screen "RIO 02 Digital Inputs" 1280x800, template "Template"
   on GenerateScreen: "TitleUpdater"()
   TextField "Text field_37" at 16,52 size 476x26; Text 'RIO #2 (Remote Inputs & Outputs Panel No. 2)'
   TextField "Text field_38" at 16,122 size 55x22; Text 'I15.0'
   TextField "Text field_39" at 16,157 size 55x22; Text 'I15.1'
   TextField "Text field_40" at 16,193 size 55x22; Text 'I15.2'
   TextField "Text field_41" at 16,229 size 55x22; Text 'I15.3'
   TextField "Text field_42" at 16,265 size 55x22; Text 'I15.4'
   TextField "Text field_43" at 16,301 size 55x22; Text 'I15.5'
   TextField "Text field_44" at 16,337 size 55x22; Text 'I15.6'
   TextField "Text field_45" at 16,373 size 55x22; Text 'I15.7'
   Circle "Circle_33" at 76,123 size 20x20
      Appearance <- "Tank 2P GTT Isolation Valve Feedback - Opened"
   Circle "Circle_34" at 76,158 size 20x20
      Appearance <- "Tank 2P GTT Isolation Valve Feedback - Closed"
   Circle "Circle_35" at 76,194 size 20x20
      Appearance <- "Tank 2P Tank Vent Valve 1 Feedback - Opened"
   Circle "Circle_36" at 76,230 size 20x20
      Appearance <- "Tank 2P Tank Vent Valve 1 Feedback - Closed"
   Circle "Circle_37" at 76,265 size 20x20
      Appearance <- "Tank 2P Tank Vent Valve 2 Feedback - Opened"
   Circle "Circle_38" at 76,301 size 20x20
      Appearance <- "Tank 2P Tank Vent Valve 2 Feedback - Closed"
   Circle "Circle_39" at 76,337 size 20x20
      Appearance <- "RIO2_SPR_DI_15_6"
   Circle "Circle_40" at 76,373 size 20x20
      Appearance <- "RIO2_SPR_DI_15_7"
   TextField "Text field_46" at 33,90 size 49x26; Text 'I0'
   TextField "Text field_47" at 16,441 size 55x22; Text 'I18.0'
   TextField "Text field_48" at 16,476 size 55x22; Text 'I18.1'
   TextField "Text field_49" at 16,512 size 55x22; Text 'I18.2'
   TextField "Text field_50" at 16,548 size 55x22; Text 'I18.3'
   TextField "Text field_51" at 16,584 size 55x22; Text 'I18.4'
   TextField "Text field_52" at 16,620 size 55x22; Text 'I18.5'
   TextField "Text field_53" at 16,656 size 55x22; Text 'I18.6'
   TextField "Text field_54" at 16,692 size 55x22; Text 'I18.7'
   Circle "Circle_41" at 76,442 size 20x20
      Appearance <- "Tank 2S GTT Isolation Valve Feedback - Opened"
   Circle "Circle_42" at 76,477 size 20x20
      Appearance <- "Tank 2S GTT Isolation Valve Feedback - Closed"
   Circle "Circle_43" at 76,513 size 20x20
      Appearance <- "Tank 2S Tank Vent Valve 1 Feedback - Opened"
   Circle "Circle_44" at 76,549 size 20x20
      Appearance <- "Tank 2S Tank Vent Valve 1 Feedback - Closed"
   Circle "Circle_45" at 76,585 size 20x20
      Appearance <- "Tank 2S Tank Vent Valve 2 Feedback - Opened"
   Circle "Circle_46" at 76,621 size 20x20
      Appearance <- "Tank 2S Tank Vent Valve 2 Feedback - Closed"
   Circle "Circle_47" at 76,657 size 20x20
      Appearance <- "RIO2_SPR_DI_18_6"
   Circle "Circle_48" at 76,693 size 20x20
      Appearance <- "RIO2_SPR_DI_18_7"
   TextField "Text field_55" at 33,409 size 49x26; Text 'I1'
   TextField "Text field_56" at 548,122 size 55x22; Text 'I21.0'
   TextField "Text field_57" at 548,157 size 55x22; Text 'I21.1'
   TextField "Text field_58" at 548,193 size 55x22; Text 'I21.2'
   TextField "Text field_59" at 548,229 size 55x22; Text 'I21.3'
   TextField "Text field_60" at 548,265 size 55x22; Text 'I21.4'
   TextField "Text field_61" at 548,301 size 55x22; Text 'I21.5'
   TextField "Text field_62" at 548,337 size 55x22; Text 'I21.6'
   TextField "Text field_63" at 548,373 size 55x22; Text 'I21.7'
   Circle "Circle_49" at 608,122 size 20x20
      Appearance <- "Tank 2P BWT Level High High Switch"
   Circle "Circle_50" at 608,157 size 20x20
      Appearance <- "RIO2 Tanks Pressure Switch Hi Hi"
   Circle "Circle_51" at 608,193 size 20x20
      Appearance <- "Tank 2S BWT Level High High Switch"
   Circle "Circle_52" at 608,229 size 20x20
      Appearance <- "RIO2_SPR_DI_21_3"
   Circle "Circle_53" at 608,265 size 20x20
      Appearance <- "RIO2_SPR_DI_21_4"
   Circle "Circle_54" at 608,301 size 20x20
      Appearance <- "RIO2_SPR_DI_21_5"
   Circle "Circle_55" at 608,337 size 20x20
      Appearance <- "RIO2_SPR_DI_21_6"
   Circle "Circle_56" at 608,373 size 20x20
      Appearance <- "RIO2_SPR_DI_21_7"
   TextField "Text field_64" at 570,90 size 49x26; Text 'I2'
   Button "HmiScreenItemData_1" at 1,1 size 150x43; TextOn 'Back'; TextOff 'Commissioning'
      on Release: ActivateScreen("Commissioning Main Page", 0)
   TextField "Text field_107" at 105,114 size 382x38; Text 'Tank 2P GTT Isolation Valve Feedback - Opened CV422'
   TextField "Text field_108" at 105,149 size 374x38; Text 'Tank 2P GTT Isolation Valve Feedback - Closed CV422'
   TextField "Text field_109" at 105,184 size 371x38; Text 'Tank 2P Tank Vent Valve 1 Feedback - Opened CV441-2P1'
   TextField "Text field_110" at 105,220 size 363x38; Text 'Tank 2P Tank Vent Valve 1 Feedback - Closed CV441-2P1'
   TextField "Text field_111" at 105,255 size 371x38; Text 'Tank 2P Tank Vent Valve 2 Feedback - Opened CV441-2P2'
   TextField "Text field_112" at 105,291 size 363x38; Text 'Tank 2P Tank Vent Valve 2 Feedback - Closed CV441-2P2'
   TextField "Text field_113" at 104,328 size 100x21; Text 'Spare Input'
   TextField "Text field_114" at 104,365 size 100x21; Text 'Spare Input'
   TextField "Text field_116" at 102,429 size 382x38; Text 'Tank 2S GTT Isolation Valve Feedback - Opened CV421-2S'
   TextField "Text field_117" at 102,465 size 374x38; Text 'Tank 2S GTT Isolation Valve Feedback - Closed CV421-2S'
   TextField "Text field_118" at 102,501 size 371x38; Text 'Tank 2S Tank Vent Valve 1 Feedback - Opened CV440-2SA'
   TextField "Text field_119" at 102,537 size 363x38; Text 'Tank 2S Tank Vent Valve 1 Feedback - Closed CV440-2SA'
   TextField "Text field_120" at 102,573 size 371x38; Text 'Tank 2S Tank Vent Valve 2 Feedback - Opened CV440-2SB'
   TextField "Text field_121" at 102,609 size 363x38; Text 'Tank 2S Tank Vent Valve 2 Feedback - Closed CV440-2SB'
   TextField "Text field_122" at 102,690 size 100x21; Text 'Spare Input'
   TextField "Text field_123" at 636,113 size 294x38; Text 'Tank 2P BWT Level High High Switch LS425-2P'
   TextField "Text field_124" at 636,148 size 270x38; Text 'RIO2 Tanks Pressure Switch Hi Hi PS436-2P/2S'
   TextField "Text field_125" at 636,184 size 294x38; Text 'Tank 2S BWT Level High High Switch LS422-2S'
   TextField "Text field_126" at 636,219 size 100x21; Text 'Spare Input'
   TextField "Text field_127" at 636,255 size 100x21; Text 'Spare Input'
   TextField "Text field_128" at 636,291 size 100x21; Text 'Spare Input'
   TextField "Text field_129" at 636,328 size 100x21; Text 'Spare Input'
   TextField "Text field_130" at 636,366 size 100x21; Text 'Spare Input'
   TextField "Text field_115" at 102,654 size 100x21; Text 'Spare Input'
   AlarmView "Alarm view_1" at 0,777 size 1280x23
   Group "Group" at 455,41 size 373x50
   Button "HmiScreenItemData_8" at 469,45 size 355x40; TextOn 'Back'; TextOff 'Text'
      on Click: "TitleUpdater"()
   TextField "Screen title" at 455,41 size 373x50; Text 'Screen title'

screen "RIO 03 Digital Inputs" 1280x800, template "Template"
   on GenerateScreen: "TitleUpdater"()
   TextField "Text field_37" at 16,52 size 476x26; Text 'RIO #3 (Remote Inputs & Outputs Panel No. 3)'
   TextField "Text field_38" at 16,122 size 55x22; Text 'I27.0'
   TextField "Text field_39" at 16,157 size 55x22; Text 'I27.1'
   TextField "Text field_40" at 16,193 size 55x22; Text 'I27.2'
   TextField "Text field_41" at 16,229 size 55x22; Text 'I27.3'
   TextField "Text field_42" at 16,265 size 55x22; Text 'I27.4'
   TextField "Text field_43" at 16,301 size 55x22; Text 'I27.5'
   TextField "Text field_44" at 16,337 size 55x22; Text 'I27.6'
   TextField "Text field_45" at 16,373 size 55x22; Text 'I27.7'
   Circle "Circle_33" at 76,123 size 20x20
      Appearance <- "Tank 3P GTT Isolation Valve Feedback - Opened"
   Circle "Circle_34" at 76,158 size 20x20
      Appearance <- "Tank 3P GTT Isolation Valve Feedback - Closed"
   Circle "Circle_35" at 76,194 size 20x20
      Appearance <- "Tank 3P Tank Vent Valve 1 Feedback - Opened"
   Circle "Circle_36" at 76,230 size 20x20
      Appearance <- "Tank 3P Tank Vent Valve 1 Feedback - Closed"
   Circle "Circle_37" at 76,265 size 20x20
      Appearance <- "Tank 3P Tank Vent Valve 2 Feedback - Opened"
   Circle "Circle_38" at 76,301 size 20x20
      Appearance <- "Tank 3P Tank Vent Valve 2 Feedback - Closed"
   Circle "Circle_39" at 76,337 size 20x20
      Appearance <- "RIO3_SPR_DI_27_6"
   Circle "Circle_40" at 76,373 size 20x20
      Appearance <- "RIO3_SPR_DI_27_7"
   TextField "Text field_46" at 33,90 size 49x26; Text 'I0'
   TextField "Text field_47" at 16,441 size 55x22; Text 'I30.0'
   TextField "Text field_48" at 16,476 size 55x22; Text 'I30.1'
   TextField "Text field_49" at 16,512 size 55x22; Text 'I30.2'
   TextField "Text field_50" at 16,548 size 55x22; Text 'I30.3'
   TextField "Text field_51" at 16,584 size 55x22; Text 'I30.4'
   TextField "Text field_52" at 16,620 size 55x22; Text 'I30.5'
   TextField "Text field_53" at 16,656 size 55x22; Text 'I30.6'
   TextField "Text field_54" at 16,692 size 55x22; Text 'I30.7'
   Circle "Circle_41" at 76,442 size 20x20
      Appearance <- "Tank 3S GTT Isolation Valve Feedback - Opened"
   Circle "Circle_42" at 76,477 size 20x20
      Appearance <- "Tank 3S GTT Isolation Valve Feedback - Closed"
   Circle "Circle_43" at 76,513 size 20x20
      Appearance <- "Tank 3S Tank Vent Valve 1 Feedback - Opened"
   Circle "Circle_44" at 76,549 size 20x20
      Appearance <- "Tank 3S Tank Vent Valve 1 Feedback - Closed"
   Circle "Circle_45" at 76,585 size 20x20
      Appearance <- "Tank 3S Tank Vent Valve 2 Feedback - Opened"
   Circle "Circle_46" at 76,621 size 20x20
      Appearance <- "Tank 3S Tank Vent Valve 2 Feedback - Closed"
   Circle "Circle_47" at 76,657 size 20x20
      Appearance <- "RIO3_SPR_DI_30_6"
   Circle "Circle_48" at 76,693 size 20x20
      Appearance <- "RIO3_SPR_DI_30_7"
   TextField "Text field_55" at 33,409 size 49x26; Text 'I1'
   TextField "Text field_56" at 548,122 size 55x22; Text 'I33.0'
   TextField "Text field_57" at 548,157 size 55x22; Text 'I33.1'
   TextField "Text field_58" at 548,193 size 55x22; Text 'I33.2'
   TextField "Text field_59" at 548,229 size 55x22; Text 'I33.3'
   TextField "Text field_60" at 548,265 size 55x22; Text 'I33.4'
   TextField "Text field_61" at 548,301 size 55x22; Text 'I33.5'
   TextField "Text field_62" at 548,337 size 55x22; Text 'I33.6'
   TextField "Text field_63" at 548,373 size 55x22; Text 'I33.7'
   Circle "Circle_49" at 608,122 size 20x20
      Appearance <- "Tank 3P BWT Level High High Switch"
   Circle "Circle_50" at 608,157 size 20x20
      Appearance <- "RIO3 Tanks Pressure Switch Hi Hi"
   Circle "Circle_51" at 608,193 size 20x20
      Appearance <- "Tank 3S BWT Level High High Switch"
   Circle "Circle_52" at 608,229 size 20x20
      Appearance <- "RIO3_SPR_DI_33_3"
   Circle "Circle_53" at 608,265 size 20x20
      Appearance <- "RIO3_SPR_DI_33_4"
   Circle "Circle_54" at 608,301 size 20x20
      Appearance <- "RIO3_SPR_DI_33_5"
   Circle "Circle_55" at 608,337 size 20x20
      Appearance <- "RIO3_SPR_DI_33_6"
   Circle "Circle_56" at 608,373 size 20x20
      Appearance <- "RIO3_SPR_DI_33_7"
   TextField "Text field_64" at 570,90 size 49x26; Text 'I2'
   Button "HmiScreenItemData_1" at 1,1 size 150x43; TextOn 'Back'; TextOff 'Commissioning'
      on Release: ActivateScreen("Commissioning Main Page", 0)
   TextField "Text field_107" at 105,114 size 382x38; Text 'Tank 3P GTT Isolation Valve Feedback - Opened CV422'
   TextField "Text field_108" at 105,149 size 374x38; Text 'Tank 3P GTT Isolation Valve Feedback - Closed CV422'
   TextField "Text field_109" at 105,184 size 371x38; Text 'Tank 3P Tank Vent Valve 1 Feedback - Opened CV441-3P1'
   TextField "Text field_110" at 105,220 size 363x38; Text 'Tank 3P Tank Vent Valve 1 Feedback - Closed CV441-3P1'
   TextField "Text field_111" at 105,255 size 371x38; Text 'Tank 3P Tank Vent Valve 2 Feedback - Opened CV441-3P2'
   TextField "Text field_112" at 105,291 size 363x38; Text 'Tank 3P Tank Vent Valve 2 Feedback - Closed CV441-3P2'
   TextField "Text field_113" at 104,328 size 100x21; Text 'Spare Input'
   TextField "Text field_114" at 104,365 size 100x21; Text 'Spare Input'
   TextField "Text field_116" at 102,429 size 382x38; Text 'Tank 3S GTT Isolation Valve Feedback - Opened CV421-3S'
   TextField "Text field_117" at 102,465 size 374x38; Text 'Tank 3S GTT Isolation Valve Feedback - Closed CV421-3S'
   TextField "Text field_118" at 102,501 size 371x38; Text 'Tank 3S Tank Vent Valve 1 Feedback - Opened CV440-3SA'
   TextField "Text field_119" at 102,537 size 363x38; Text 'Tank 3S Tank Vent Valve 1 Feedback - Closed CV440-3SA'
   TextField "Text field_120" at 102,573 size 371x38; Text 'Tank 3S Tank Vent Valve 2 Feedback - Opened CV440-3SB'
   TextField "Text field_121" at 102,609 size 363x38; Text 'Tank 3S Tank Vent Valve 2 Feedback - Closed CV440-3SB'
   TextField "Text field_122" at 102,690 size 100x21; Text 'Spare Input'
   TextField "Text field_123" at 636,113 size 294x38; Text 'Tank 3P BWT Level High High Switch LS425-3P'
   TextField "Text field_124" at 636,148 size 270x38; Text 'RIO3 Tanks Pressure Switch Hi Hi PS436-3P/3S'
   TextField "Text field_125" at 636,184 size 294x38; Text 'Tank 3S BWT Level High High Switch LS422-3S'
   TextField "Text field_126" at 636,219 size 100x21; Text 'Spare Input'
   TextField "Text field_127" at 636,255 size 100x21; Text 'Spare Input'
   TextField "Text field_128" at 636,291 size 100x21; Text 'Spare Input'
   TextField "Text field_129" at 636,328 size 100x21; Text 'Spare Input'
   TextField "Text field_130" at 636,366 size 100x21; Text 'Spare Input'
   TextField "Text field_115" at 102,654 size 100x21; Text 'Spare Input'
   AlarmView "Alarm view_1" at 0,777 size 1280x23
   Group "Group" at 455,41 size 373x50
   Button "HmiScreenItemData_8" at 469,45 size 355x40; TextOn 'Back'; TextOff 'Text'
      on Click: "TitleUpdater"()
   TextField "Screen title" at 455,41 size 373x50; Text 'Screen title'

screen "RIO 04 Digital Inputs" 1280x800, template "Template"
   on GenerateScreen: "TitleUpdater"()
   TextField "Text field_37" at 16,52 size 476x26; Text 'RIO #4 (Remote Inputs & Outputs Panel No. 4)'
   TextField "Text field_38" at 16,122 size 55x22; Text 'I39.0'
   TextField "Text field_39" at 16,157 size 55x22; Text 'I39.1'
   TextField "Text field_40" at 16,193 size 55x22; Text 'I39.2'
   TextField "Text field_41" at 16,229 size 55x22; Text 'I39.3'
   TextField "Text field_42" at 16,265 size 55x22; Text 'I39.4'
   TextField "Text field_43" at 16,301 size 55x22; Text 'I39.5'
   TextField "Text field_44" at 16,337 size 55x22; Text 'I39.6'
   TextField "Text field_45" at 16,373 size 55x22; Text 'I39.7'
   Circle "Circle_33" at 76,123 size 20x20
      Appearance <- "Tank 4P GTT Isolation Valve Feedback - Opened"
   Circle "Circle_34" at 76,158 size 20x20
      Appearance <- "Tank 4P GTT Isolation Valve Feedback - Closed"
   Circle "Circle_35" at 76,194 size 20x20
      Appearance <- "Tank 4P Tank Vent Valve 1 Feedback - Opened"
   Circle "Circle_36" at 76,230 size 20x20
      Appearance <- "Tank 4P Tank Vent Valve 1 Feedback - Closed"
   Circle "Circle_37" at 76,265 size 20x20
      Appearance <- "Tank 4P Tank Vent Valve 2 Feedback - Opened"
   Circle "Circle_38" at 76,301 size 20x20
      Appearance <- "Tank 4P Tank Vent Valve 2 Feedback - Closed"
   Circle "Circle_39" at 76,337 size 20x20
      Appearance <- "RIO4_SPR_DI_139_6"
   Circle "Circle_40" at 76,373 size 20x20
      Appearance <- "RIO4_SPR_DI_139_7"
   TextField "Text field_46" at 33,90 size 49x26; Text 'I0'
   TextField "Text field_47" at 16,441 size 55x22; Text 'I42.0'
   TextField "Text field_48" at 16,476 size 55x22; Text 'I42.1'
   TextField "Text field_49" at 16,512 size 55x22; Text 'I42.2'
   TextField "Text field_50" at 16,548 size 55x22; Text 'I42.3'
   TextField "Text field_51" at 16,584 size 55x22; Text 'I42.4'
   TextField "Text field_52" at 16,620 size 55x22; Text 'I42.5'
   TextField "Text field_53" at 16,656 size 55x22; Text 'I42.6'
   TextField "Text field_54" at 16,692 size 55x22; Text 'I42.7'
   Circle "Circle_41" at 76,442 size 20x20
      Appearance <- "Tank 4S GTT Isolation Valve Feedback - Opened"
   Circle "Circle_42" at 76,477 size 20x20
      Appearance <- "Tank 4S GTT Isolation Valve Feedback - Closed"
   Circle "Circle_43" at 76,513 size 20x20
      Appearance <- "Tank 4S Tank Vent Valve 1 Feedback - Opened"
   Circle "Circle_44" at 76,549 size 20x20
      Appearance <- "Tank 4S Tank Vent Valve 1 Feedback - Closed"
   Circle "Circle_45" at 76,585 size 20x20
      Appearance <- "Tank 4S Tank Vent Valve 2 Feedback - Opened"
   Circle "Circle_46" at 76,621 size 20x20
      Appearance <- "Tank 4S Tank Vent Valve 2 Feedback - Closed"
   Circle "Circle_47" at 76,657 size 20x20
      Appearance <- "RIO4_SPR_DI_142_6"
   Circle "Circle_48" at 76,693 size 20x20
      Appearance <- "RIO4_SPR_DI_142_7"
   TextField "Text field_55" at 33,409 size 49x26; Text 'I1'
   TextField "Text field_56" at 548,122 size 55x22; Text 'I45.0'
   TextField "Text field_57" at 548,157 size 55x22; Text 'I45.1'
   TextField "Text field_58" at 548,193 size 55x22; Text 'I45.2'
   TextField "Text field_59" at 548,229 size 55x22; Text 'I45.3'
   TextField "Text field_60" at 548,265 size 55x22; Text 'I45.4'
   TextField "Text field_61" at 548,301 size 55x22; Text 'I45.5'
   TextField "Text field_62" at 548,337 size 55x22; Text 'I45.6'
   TextField "Text field_63" at 548,373 size 55x22; Text 'I45.7'
   Circle "Circle_49" at 608,122 size 20x20
      Appearance <- "Tank 4P BWT Level High High Switch"
   Circle "Circle_50" at 608,157 size 20x20
      Appearance <- "RIO4 Tanks Pressure Switch Hi Hi"
   Circle "Circle_51" at 608,193 size 20x20
      Appearance <- "Tank 4S BWT Level High High Switch"
   Circle "Circle_52" at 608,229 size 20x20
      Appearance <- "RIO4_SPR_DI_145_3"
   Circle "Circle_53" at 608,265 size 20x20
      Appearance <- "RIO4_SPR_DI_145_4"
   Circle "Circle_54" at 608,301 size 20x20
      Appearance <- "RIO4_SPR_DI_145_5"
   Circle "Circle_55" at 608,337 size 20x20
      Appearance <- "RIO4_SPR_DI_145_6"
   Circle "Circle_56" at 608,373 size 20x20
      Appearance <- "RIO4_SPR_DI_145_7"
   TextField "Text field_64" at 570,90 size 49x26; Text 'I2'
   Button "HmiScreenItemData_1" at 1,1 size 150x43; TextOn 'Back'; TextOff 'Commissioning'
      on Release: ActivateScreen("Commissioning Main Page", 0)
   TextField "Text field_107" at 105,114 size 382x38; Text 'Tank 4P GTT Isolation Valve Feedback - Opened CV422'
   TextField "Text field_108" at 105,149 size 374x38; Text 'Tank 4P GTT Isolation Valve Feedback - Closed CV422'
   TextField "Text field_109" at 105,184 size 371x38; Text 'Tank 4P Tank Vent Valve 1 Feedback - Opened CV441-4P1'
   TextField "Text field_110" at 105,220 size 363x38; Text 'Tank 4P Tank Vent Valve 1 Feedback - Closed CV441-4P1'
   TextField "Text field_111" at 105,255 size 371x38; Text 'Tank 4P Tank Vent Valve 2 Feedback - Opened CV441-4P2'
   TextField "Text field_112" at 105,291 size 363x38; Text 'Tank 4P Tank Vent Valve 2 Feedback - Closed CV441-4P2'
   TextField "Text field_113" at 104,328 size 100x21; Text 'Spare Input'
   TextField "Text field_114" at 104,365 size 100x21; Text 'Spare Input'
   TextField "Text field_116" at 102,429 size 382x38; Text 'Tank 4S GTT Isolation Valve Feedback - Opened CV421-4S'
   TextField "Text field_117" at 102,465 size 374x38; Text 'Tank 4S GTT Isolation Valve Feedback - Closed CV421-4S'
   TextField "Text field_118" at 102,501 size 371x38; Text 'Tank 4S Tank Vent Valve 1 Feedback - Opened CV440-4SA'
   TextField "Text field_119" at 102,537 size 363x38; Text 'Tank 4S Tank Vent Valve 1 Feedback - Closed CV440-4SA'
   TextField "Text field_120" at 102,573 size 371x38; Text 'Tank 4S Tank Vent Valve 2 Feedback - Opened CV440-4SB'
   TextField "Text field_121" at 102,609 size 363x38; Text 'Tank 4S Tank Vent Valve 2 Feedback - Closed CV440-4SB'
   TextField "Text field_122" at 102,690 size 100x21; Text 'Spare Input'
   TextField "Text field_123" at 636,113 size 294x38; Text 'Tank 4P BWT Level High High Switch LS425-4P'
   TextField "Text field_124" at 636,148 size 270x38; Text 'RIO4 Tanks Pressure Switch Hi Hi PS436-4P/4S'
   TextField "Text field_125" at 636,184 size 294x38; Text 'Tank 4S BWT Level High High Switch LS422-4S'
   TextField "Text field_126" at 636,219 size 100x21; Text 'Spare Input'
   TextField "Text field_127" at 636,255 size 100x21; Text 'Spare Input'
   TextField "Text field_128" at 636,291 size 100x21; Text 'Spare Input'
   TextField "Text field_129" at 636,328 size 100x21; Text 'Spare Input'
   TextField "Text field_130" at 636,366 size 100x21; Text 'Spare Input'
   TextField "Text field_115" at 102,654 size 100x21; Text 'Spare Input'
   AlarmView "Alarm view_1" at 0,777 size 1280x23
   Group "Group" at 455,41 size 373x50
   Button "HmiScreenItemData_8" at 469,45 size 355x40; TextOn 'Back'; TextOff 'Text'
      on Click: "TitleUpdater"()
   TextField "Screen title" at 455,41 size 373x50; Text 'Screen title'

screen "RIO 05 Digital Inputs" 1280x800, template "Template"
   on GenerateScreen: "TitleUpdater"()
   TextField "Text field_37" at 16,52 size 476x26; Text 'RIO #5 (Remote Inputs & Outputs Panel No. 5)'
   TextField "Text field_38" at 16,122 size 55x22; Text 'I51.0'
   TextField "Text field_39" at 16,157 size 55x22; Text 'I51.1'
   TextField "Text field_40" at 16,193 size 55x22; Text 'I51.2'
   TextField "Text field_41" at 16,229 size 55x22; Text 'I51.3'
   TextField "Text field_42" at 16,265 size 55x22; Text 'I51.4'
   TextField "Text field_43" at 16,301 size 55x22; Text 'I51.5'
   TextField "Text field_44" at 16,337 size 55x22; Text 'I51.6'
   TextField "Text field_45" at 16,373 size 55x22; Text 'I51.7'
   Circle "Circle_33" at 76,123 size 20x20
      Appearance <- "Tank 5P GTT Isolation Valve Feedback - Opened"
   Circle "Circle_34" at 76,158 size 20x20
      Appearance <- "Tank 5P GTT Isolation Valve Feedback - Closed"
   Circle "Circle_35" at 76,194 size 20x20
      Appearance <- "Tank 5P Tank Vent Valve 1 Feedback - Opened"
   Circle "Circle_36" at 76,230 size 20x20
      Appearance <- "Tank 5P Tank Vent Valve 1 Feedback - Closed"
   Circle "Circle_37" at 76,265 size 20x20
      Appearance <- "Tank 5P Tank Vent Valve 2 Feedback - Opened"
   Circle "Circle_38" at 76,301 size 20x20
      Appearance <- "Tank 5P Tank Vent Valve 2 Feedback - Closed"
   Circle "Circle_39" at 76,337 size 20x20
      Appearance <- "RIO5_SPR_DI_51_6"
   Circle "Circle_40" at 76,373 size 20x20
      Appearance <- "RIO5_SPR_DI_51_7"
   TextField "Text field_46" at 33,90 size 49x26; Text 'I0'
   TextField "Text field_47" at 16,441 size 55x22; Text 'I54.0'
   TextField "Text field_48" at 16,476 size 55x22; Text 'I54.1'
   TextField "Text field_49" at 16,512 size 55x22; Text 'I54.2'
   TextField "Text field_50" at 16,548 size 55x22; Text 'I54.3'
   TextField "Text field_51" at 16,584 size 55x22; Text 'I54.4'
   TextField "Text field_52" at 16,620 size 55x22; Text 'I54.5'
   TextField "Text field_53" at 16,656 size 55x22; Text 'I54.6'
   TextField "Text field_54" at 16,692 size 55x22; Text 'I54.7'
   Circle "Circle_41" at 76,442 size 20x20
      Appearance <- "Tank 5S GTT Isolation Valve Feedback - Opened"
   Circle "Circle_42" at 76,477 size 20x20
      Appearance <- "Tank 5S GTT Isolation Valve Feedback - Closed"
   Circle "Circle_43" at 76,513 size 20x20
      Appearance <- "Tank 5S Tank Vent Valve 1 Feedback - Opened"
   Circle "Circle_44" at 76,549 size 20x20
      Appearance <- "Tank 5S Tank Vent Valve 1 Feedback - Closed"
   Circle "Circle_45" at 76,585 size 20x20
      Appearance <- "Tank 5S Tank Vent Valve 2 Feedback - Opened"
   Circle "Circle_46" at 76,621 size 20x20
      Appearance <- "Tank 5S Tank Vent Valve 2 Feedback - Closed"
   Circle "Circle_47" at 76,657 size 20x20
      Appearance <- "RIO5_SPR_DI_54_6"
   Circle "Circle_48" at 76,693 size 20x20
      Appearance <- "RIO5_SPR_DI_54_7"
   TextField "Text field_55" at 33,409 size 49x26; Text 'I1'
   TextField "Text field_56" at 548,122 size 55x22; Text 'I57.0'
   TextField "Text field_57" at 548,157 size 55x22; Text 'I57.1'
   TextField "Text field_58" at 548,193 size 55x22; Text 'I57.2'
   TextField "Text field_59" at 548,229 size 55x22; Text 'I57.3'
   TextField "Text field_60" at 548,265 size 55x22; Text 'I57.4'
   TextField "Text field_61" at 548,301 size 55x22; Text 'I57.5'
   TextField "Text field_62" at 548,337 size 55x22; Text 'I57.6'
   TextField "Text field_63" at 548,373 size 55x22; Text 'I57.7'
   Circle "Circle_49" at 608,122 size 20x20
      Appearance <- "Tank 5P BWT Level High High Switch"
   Circle "Circle_50" at 608,157 size 20x20
      Appearance <- "RIO5 Tanks Pressure Switch Hi Hi"
   Circle "Circle_51" at 608,193 size 20x20
      Appearance <- "Tank 5S BWT Level High High Switch"
   Circle "Circle_52" at 608,229 size 20x20
      Appearance <- "RIO5_SPR_DI_57_3"
   Circle "Circle_53" at 608,265 size 20x20
      Appearance <- "RIO5_SPR_DI_57_4"
   Circle "Circle_54" at 608,301 size 20x20
      Appearance <- "RIO5_SPR_DI_57_5"
   Circle "Circle_55" at 608,337 size 20x20
      Appearance <- "RIO5_SPR_DI_57_6"
   Circle "Circle_56" at 608,373 size 20x20
      Appearance <- "RIO5_SPR_DI_57_7"
   TextField "Text field_64" at 570,90 size 49x26; Text 'I2'
   Button "HmiScreenItemData_1" at 1,1 size 150x43; TextOn 'Back'; TextOff 'Commissioning'
      on Release: ActivateScreen("Commissioning Main Page", 0)
   TextField "Text field_107" at 105,114 size 382x38; Text 'Tank 5P GTT Isolation Valve Feedback - Opened CV422'
   TextField "Text field_108" at 105,149 size 374x38; Text 'Tank 5P GTT Isolation Valve Feedback - Closed CV422'
   TextField "Text field_109" at 105,184 size 371x38; Text 'Tank 5P Tank Vent Valve 1 Feedback - Opened CV441-5P1'
   TextField "Text field_110" at 105,220 size 363x38; Text 'Tank 5P Tank Vent Valve 1 Feedback - Closed CV441-5P1'
   TextField "Text field_111" at 105,255 size 371x38; Text 'Tank 5P Tank Vent Valve 2 Feedback - Opened CV441-5P2'
   TextField "Text field_112" at 105,291 size 363x38; Text 'Tank 5P Tank Vent Valve 2 Feedback - Closed CV441-5P2'
   TextField "Text field_113" at 104,328 size 100x21; Text 'Spare Input'
   TextField "Text field_114" at 104,365 size 100x21; Text 'Spare Input'
   TextField "Text field_116" at 102,429 size 382x38; Text 'Tank 5S GTT Isolation Valve Feedback - Opened CV421-5S'
   TextField "Text field_117" at 102,465 size 374x38; Text 'Tank 5S GTT Isolation Valve Feedback - Closed CV421-5S'
   TextField "Text field_118" at 102,501 size 371x38; Text 'Tank 5S Tank Vent Valve 1 Feedback - Opened CV440-5SA'
   TextField "Text field_119" at 102,537 size 363x38; Text 'Tank 5S Tank Vent Valve 1 Feedback - Closed CV440-5SA'
   TextField "Text field_120" at 102,573 size 371x38; Text 'Tank 5S Tank Vent Valve 2 Feedback - Opened CV440-5SB'
   TextField "Text field_121" at 102,609 size 363x38; Text 'Tank 5S Tank Vent Valve 2 Feedback - Closed CV440-5SB'
   TextField "Text field_122" at 102,690 size 100x21; Text 'Spare Input'
   TextField "Text field_123" at 636,113 size 294x38; Text 'Tank 5P BWT Level High High Switch LS425-5P'
   TextField "Text field_124" at 636,148 size 270x38; Text 'RIO5 Tanks Pressure Switch Hi Hi PS436-5P/5S'
   TextField "Text field_125" at 636,184 size 294x38; Text 'Tank 5S BWT Level High High Switch LS422-5S'
   TextField "Text field_126" at 636,219 size 100x21; Text 'Spare Input'
   TextField "Text field_127" at 636,255 size 100x21; Text 'Spare Input'
   TextField "Text field_128" at 636,291 size 100x21; Text 'Spare Input'
   TextField "Text field_129" at 636,328 size 100x21; Text 'Spare Input'
   TextField "Text field_130" at 636,366 size 100x21; Text 'Spare Input'
   TextField "Text field_115" at 102,654 size 100x21; Text 'Spare Input'
   AlarmView "Alarm view_1" at 0,777 size 1280x23
   Group "Group" at 455,41 size 373x50
   Button "HmiScreenItemData_8" at 469,45 size 355x40; TextOn 'Back'; TextOff 'Text'
      on Click: "TitleUpdater"()
   TextField "Screen title" at 455,41 size 373x50; Text 'Screen title'

screen "RIO 06 Digital Inputs" 1280x800, template "Template"
   on GenerateScreen: "TitleUpdater"()
   TextField "Text field_37" at 16,52 size 476x26; Text 'RIO #6 (Remote Inputs & Outputs Panel No. 6)'
   TextField "Text field_38" at 16,122 size 55x22; Text 'I60.0'
   TextField "Text field_39" at 16,157 size 55x22; Text 'I60.1'
   TextField "Text field_40" at 16,193 size 55x22; Text 'I60.2'
   TextField "Text field_41" at 16,229 size 55x22; Text 'I60.3'
   TextField "Text field_42" at 16,265 size 55x22; Text 'I60.4'
   TextField "Text field_43" at 16,301 size 55x22; Text 'I60.5'
   TextField "Text field_44" at 16,337 size 55x22; Text 'I60.6'
   TextField "Text field_45" at 16,373 size 55x22; Text 'I60.7'
   Circle "Circle_33" at 76,123 size 20x20
      Appearance <- "Tank 6P GTT Isolation Valve Feedback - Opened"
   Circle "Circle_34" at 76,158 size 20x20
      Appearance <- "Tank 6P GTT Isolation Valve Feedback - Closed"
   Circle "Circle_35" at 76,194 size 20x20
      Appearance <- "Tank 6P Tank Vent Valve 1 Feedback - Opened"
   Circle "Circle_36" at 76,230 size 20x20
      Appearance <- "Tank 6P Tank Vent Valve 1 Feedback - Closed"
   Circle "Circle_37" at 76,265 size 20x20
      Appearance <- "Tank 6P Tank Vent Valve 2 Feedback - Opened"
   Circle "Circle_38" at 76,301 size 20x20
      Appearance <- "Tank 6P Tank Vent Valve 2 Feedback - Closed"
   Circle "Circle_39" at 76,337 size 20x20
      Appearance <- "RIO6_SPR_DI_60_6"
   Circle "Circle_40" at 76,373 size 20x20
      Appearance <- "RIO6_SPR_DI_60_7"
   TextField "Text field_46" at 33,90 size 49x26; Text 'I0'
   TextField "Text field_47" at 16,441 size 55x22; Text 'I63.0'
   TextField "Text field_48" at 16,476 size 55x22; Text 'I63.1'
   TextField "Text field_49" at 16,512 size 55x22; Text 'I63.2'
   TextField "Text field_50" at 16,548 size 55x22; Text 'I63.3'
   TextField "Text field_51" at 16,584 size 55x22; Text 'I63.4'
   TextField "Text field_52" at 16,620 size 55x22; Text 'I63.5'
   TextField "Text field_53" at 16,656 size 55x22; Text 'I63.6'
   TextField "Text field_54" at 16,692 size 55x22; Text 'I63.7'
   Circle "Circle_41" at 76,442 size 20x20
      Appearance <- "Tank 6S GTT Isolation Valve Feedback - Opened"
   Circle "Circle_42" at 76,477 size 20x20
      Appearance <- "Tank 6S GTT Isolation Valve Feedback - Closed"
   Circle "Circle_43" at 76,513 size 20x20
      Appearance <- "Tank 6S Tank Vent Valve 1 Feedback - Opened"
   Circle "Circle_44" at 76,549 size 20x20
      Appearance <- "Tank 6S Tank Vent Valve 1 Feedback - Closed"
   Circle "Circle_45" at 76,585 size 20x20
      Appearance <- "Tank 6S Tank Vent Valve 2 Feedback - Opened"
   Circle "Circle_46" at 76,621 size 20x20
      Appearance <- "Tank 6S Tank Vent Valve 2 Feedback - Closed"
   Circle "Circle_47" at 76,657 size 20x20
      Appearance <- "RIO6_SPR_DI_63_6"
   Circle "Circle_48" at 76,693 size 20x20
      Appearance <- "RIO6_SPR_DI_63_7"
   TextField "Text field_55" at 33,409 size 49x26; Text 'I1'
   TextField "Text field_56" at 548,122 size 55x22; Text 'I66.0'
   TextField "Text field_57" at 548,157 size 55x22; Text 'I66.1'
   TextField "Text field_58" at 548,193 size 55x22; Text 'I66.2'
   TextField "Text field_59" at 548,229 size 55x22; Text 'I66.3'
   TextField "Text field_60" at 548,265 size 55x22; Text 'I66.4'
   TextField "Text field_61" at 548,301 size 55x22; Text 'I66.5'
   TextField "Text field_62" at 548,337 size 55x22; Text 'I66.6'
   TextField "Text field_63" at 548,373 size 55x22; Text 'I66.7'
   Circle "Circle_49" at 608,122 size 20x20
      Appearance <- "Tank 6P BWT Level High High Switch"
   Circle "Circle_50" at 608,157 size 20x20
      Appearance <- "RIO6 Tanks Pressure Switch Hi Hi"
   Circle "Circle_51" at 608,193 size 20x20
      Appearance <- "Tank 6S BWT Level High High Switch"
   Circle "Circle_52" at 608,229 size 20x20
      Appearance <- "RIO6_SPR_DI_66_3"
   Circle "Circle_53" at 608,265 size 20x20
      Appearance <- "RIO6_SPR_DI_66_4"
   Circle "Circle_54" at 608,301 size 20x20
      Appearance <- "RIO6_SPR_DI_66_5"
   Circle "Circle_55" at 608,337 size 20x20
      Appearance <- "RIO6_SPR_DI_66_6"
   Circle "Circle_56" at 608,373 size 20x20
      Appearance <- "RIO6_SPR_DI_66_7"
   TextField "Text field_64" at 570,90 size 49x26; Text 'I2'
   Button "HmiScreenItemData_1" at 1,1 size 150x43; TextOn 'Back'; TextOff 'Commissioning'
      on Release: ActivateScreen("Commissioning Main Page", 0)
   TextField "Text field_107" at 105,114 size 382x38; Text 'Tank 6P GTT Isolation Valve Feedback - Opened CV422'
   TextField "Text field_108" at 105,149 size 374x38; Text 'Tank 6P GTT Isolation Valve Feedback - Closed CV422'
   TextField "Text field_109" at 105,184 size 371x38; Text 'Tank 6P Tank Vent Valve 1 Feedback - Opened CV441-6P1'
   TextField "Text field_110" at 105,220 size 363x38; Text 'Tank 6P Tank Vent Valve 1 Feedback - Closed CV441-6P1'
   TextField "Text field_111" at 105,255 size 371x38; Text 'Tank 6P Tank Vent Valve 2 Feedback - Opened CV441-6P2'
   TextField "Text field_112" at 105,291 size 363x38; Text 'Tank 6P Tank Vent Valve 2 Feedback - Closed CV441-6P2'
   TextField "Text field_113" at 104,328 size 100x21; Text 'Spare Input'
   TextField "Text field_114" at 104,365 size 100x21; Text 'Spare Input'
   TextField "Text field_116" at 102,429 size 382x38; Text 'Tank 6S GTT Isolation Valve Feedback - Opened CV421-6S'
   TextField "Text field_117" at 102,465 size 374x38; Text 'Tank 6S GTT Isolation Valve Feedback - Closed CV421-6S'
   TextField "Text field_118" at 102,501 size 371x38; Text 'Tank 6S Tank Vent Valve 1 Feedback - Opened CV440-6SA'
   TextField "Text field_119" at 102,537 size 363x38; Text 'Tank 6S Tank Vent Valve 1 Feedback - Closed CV440-6SA'
   TextField "Text field_120" at 102,573 size 371x38; Text 'Tank 6S Tank Vent Valve 2 Feedback - Opened CV440-6SB'
   TextField "Text field_121" at 102,609 size 363x38; Text 'Tank 6S Tank Vent Valve 2 Feedback - Closed CV440-6SB'
   TextField "Text field_122" at 102,690 size 100x21; Text 'Spare Input'
   TextField "Text field_123" at 636,113 size 294x38; Text 'Tank 6P BWT Level High High Switch LS425-6P'
   TextField "Text field_124" at 636,148 size 270x38; Text 'RIO6 Tanks Pressure Switch Hi Hi PS436-6P/6S'
   TextField "Text field_125" at 636,184 size 294x38; Text 'Tank 6S BWT Level High High Switch LS422-6S'
   TextField "Text field_126" at 636,219 size 100x21; Text 'Spare Input'
   TextField "Text field_127" at 636,255 size 100x21; Text 'Spare Input'
   TextField "Text field_128" at 636,291 size 100x21; Text 'Spare Input'
   TextField "Text field_129" at 636,328 size 100x21; Text 'Spare Input'
   TextField "Text field_130" at 636,366 size 100x21; Text 'Spare Input'
   TextField "Text field_115" at 102,654 size 100x21; Text 'Spare Input'
   AlarmView "Alarm view_1" at 0,777 size 1280x23
   Group "Group" at 455,41 size 373x50
   Button "HmiScreenItemData_8" at 469,45 size 355x40; TextOn 'Back'; TextOff 'Text'
      on Click: "TitleUpdater"()
   TextField "Screen title" at 455,41 size 373x50; Text 'Screen title'

screen "RIO 07 Digital Inputs" 1280x800, template "Template"
   on GenerateScreen: "TitleUpdater"()
   TextField "Text field_37" at 16,52 size 476x26; Text 'RIO #7 (Remote Inputs & Outputs Panel No. 7)'
   TextField "Text field_38" at 16,122 size 55x22; Text 'I75.0'
   TextField "Text field_39" at 16,157 size 55x22; Text 'I75.1'
   TextField "Text field_40" at 16,193 size 55x22; Text 'I75.2'
   TextField "Text field_41" at 16,229 size 55x22; Text 'I75.3'
   TextField "Text field_42" at 16,265 size 55x22; Text 'I75.4'
   TextField "Text field_43" at 16,301 size 55x22; Text 'I75.5'
   TextField "Text field_44" at 16,337 size 55x22; Text 'I75.6'
   TextField "Text field_45" at 16,373 size 55x22; Text 'I75.7'
   Circle "Circle_33" at 76,123 size 20x20
      Appearance <- "APT GTT Isolation Valve Feedback - Opened"
   Circle "Circle_34" at 76,158 size 20x20
      Appearance <- "APT GTT Isolation Valve Feedback - Closed"
   Circle "Circle_35" at 76,194 size 20x20
      Appearance <- "APT Tank Vent Valve 1 Feedback - Opened"
   Circle "Circle_36" at 76,230 size 20x20
      Appearance <- "APT Tank Vent Valve 1 Feedback - Closed"
   Circle "Circle_37" at 76,265 size 20x20
      Appearance <- "APT Tank Vent Valve 2 Feedback - Opened"
   Circle "Circle_38" at 76,301 size 20x20
      Appearance <- "APT Tank Vent Valve 2 Feedback - Closed"
   Circle "Circle_39" at 76,337 size 20x20
      Appearance <- "RIO7_SPR_DI_175_6"
   Circle "Circle_40" at 76,373 size 20x20
      Appearance <- "RIO7_SPR_DI_175_7"
   TextField "Text field_46" at 33,90 size 49x26; Text 'I0'
   TextField "Text field_56" at 548,122 size 55x22; Text 'I78.0'
   TextField "Text field_57" at 548,157 size 55x22; Text 'I78.1'
   TextField "Text field_58" at 548,193 size 55x22; Text 'I78.2'
   TextField "Text field_59" at 548,229 size 55x22; Text 'I78.3'
   TextField "Text field_60" at 548,265 size 55x22; Text 'I78.4'
   TextField "Text field_61" at 548,301 size 55x22; Text 'I78.5'
   TextField "Text field_62" at 548,337 size 55x22; Text 'I78.6'
   TextField "Text field_63" at 548,373 size 55x22; Text 'I78.7'
   Circle "Circle_49" at 608,122 size 20x20
      Appearance <- "APT BWT Level High High Switch"
   Circle "Circle_50" at 608,157 size 20x20
      Appearance <- "RIO7 Tank Pressure Switch Hi Hi"
   Circle "Circle_51" at 608,193 size 20x20
      Appearance <- "RIO7_SPR_DI_178_2"
   Circle "Circle_52" at 608,229 size 20x20
      Appearance <- "RIO7_SPR_DI_178_3"
   Circle "Circle_53" at 608,265 size 20x20
      Appearance <- "RIO7_SPR_DI_178_4"
   Circle "Circle_54" at 608,301 size 20x20
      Appearance <- "RIO7_SPR_DI_178_5"
   Circle "Circle_55" at 608,337 size 20x20
      Appearance <- "RIO7_SPR_DI_178_6"
   Circle "Circle_56" at 608,373 size 20x20
      Appearance <- "RIO7_SPR_DI_178_7"
   TextField "Text field_64" at 570,90 size 49x26; Text 'I1'
   Button "HmiScreenItemData_1" at 1,1 size 150x43; TextOn 'Back'; TextOff 'Commissioning'
      on Release: ActivateScreen("Commissioning Main Page", 0)
   TextField "Text field_107" at 105,114 size 393x38; Text 'Tank APT GTT Isolation Valve Feedback - Opened CV422'
   TextField "Text field_108" at 105,149 size 385x38; Text 'Tank APT GTT Isolation Valve Feedback - Closed CV422'
   TextField "Text field_109" at 105,184 size 382x38; Text 'Tank APT Tank Vent Valve 1 Feedback - Opened CV441-APT1'
   TextField "Text field_110" at 105,220 size 374x38; Text 'Tank APT Tank Vent Valve 1 Feedback - Closed CV441-APT1'
   TextField "Text field_111" at 105,255 size 382x38; Text 'Tank APT Tank Vent Valve 2 Feedback - Opened CV441-APT2'
   TextField "Text field_112" at 105,291 size 374x38; Text 'Tank APT Tank Vent Valve 2 Feedback - Closed CV441-APT2'
   TextField "Text field_113" at 104,328 size 100x21; Text 'Spare Input'
   TextField "Text field_114" at 104,365 size 100x21; Text 'Spare Input'
   TextField "Text field_123" at 636,113 size 294x38; Text 'Tank APT BWT Level High High Switch LS425-APT'
   TextField "Text field_124" at 636,148 size 270x38; Text 'RIO7 Tanks Pressure Switch Hi Hi PS436-APT'
   TextField "Text field_125" at 636,184 size 100x21; Text 'Spare Input'
   TextField "Text field_126" at 636,219 size 100x21; Text 'Spare Input'
   TextField "Text field_127" at 636,255 size 100x21; Text 'Spare Input'
   TextField "Text field_128" at 636,291 size 100x21; Text 'Spare Input'
   TextField "Text field_129" at 636,328 size 100x21; Text 'Spare Input'
   TextField "Text field_130" at 636,366 size 100x21; Text 'Spare Input'
   AlarmView "Alarm view_1" at 0,777 size 1280x23
   Group "Group" at 455,41 size 373x50
   Button "HmiScreenItemData_8" at 469,45 size 355x40; TextOn 'Back'; TextOff 'Text'
      on Click: "TitleUpdater"()
   TextField "Screen title" at 455,41 size 373x50; Text 'Screen title'

PopupScreen "BWT Mode Warning" 665x250
   Button "Button_1" at 0,0 size 665x250; TextOff 'BWT Mode Not Selected. Select BWT Mode for Tank Treatment. For Cargo Blanketing use IGG Controls.'
      on Release: ActivateScreen("Balast Water Treatment Setup", 0)
   Button "Button_2" at 208,187 size 250x35; TextOff 'OK, Select Treatment Mode'
      on Release: ActivateScreen("Balast Water Treatment Setup", 0); function_efd93a16("BWT Mode Warning", 0, 0, -1, -1, 1)

PopupScreen "IGG Temperature Trends" 810x675
   on GenerateScreen: "TitleUpdater"()
   Button "Button_1" at 753,0 size 56x38; TextOff 'Text'; PictureOff "Graphic_286"
      on Click: function_efd93a16("IGG Temperature Trends", 0, 0, -1, -1, 1)
   GraphicView "Graphic view_2" at 2,2 size 751x35; Picture "Graphic_287"
   TrendView "Trend view_1" at 1,40 size 805x635
      Visibility <- "80_From_HMI_BWT_BYPASS"
      ValueAxis2End <- "84_Setpoints_PIT359_HighHigh"
      ValueAxis2Begin <- "84_Setpoints_PIT359_LowLow"
   TextField "Text field_1" at 282,7 size 252x26; Text 'IGG Temperature Trends'

screen "Reports" 1280x800, template "Template"
   RecipeView "Recipe view_1" at 854,43 size 400x350; Tag4RecipeNumber "Recipe Tag"; Tag4DataRecord "Record Data Tag"
   Button "HmiScreenItemData_1" at 2,2 size 159x51; TextOn 'Back'; TextOff 'Home'
      on Release: ActivateScreen("01 Home", 0)

screen "Balast Water Treatment Plant Tank Levels" 1280x800, template "Template"
   on GenerateScreen: "User_Change"(); "TitleUpdater"()
   Button "HmiScreenItemData_1" at 1,1 size 150x40; TextOn 'Back'; TextOff 'Main Index'
      on Release: ActivateScreen("02 Main Index", 0)
   TextField "Text field_63" at 383,107 size 72x30; Text 'Pre Dwell Time'
   Circle "Circle_29" at 1047,85 size 20x20
      Appearance <- "2102_TIME_CALCS_DB_POST_DWELL_TMR_DN"
   Button "HmiScreenItemData_9" at 10,60 size 158x27; TextOn 'Back'; TextOff 'BWTS Control'
   Button "HmiScreenItemData_4" at 14,150 size 75x47; TextOn 'Back'; TextOff 'Stop'; Authorization "Operate"
      on Release: function_efd93a16("BWTS Stop Confirm", 400, 200, -1, -1, 1)
      ObjectEnable <- "82_To_HMI_CRNT_MODE_GCU"
   Circle "Circle_20" at 137,105 size 29x29
      Appearance <- "80_From_HMI_RUN_IGG(1)"
   Button "HmiScreenItemData_3" at 14,93 size 75x47; TextOn 'Back'; TextOff 'Start'; Authorization "Operate"
      on Release: function_efd93a16("BWTS Start Confirm", 400, 200, -1, -1, 1)
      ObjectEnable <- "82_To_HMI_CRNT_MODE_GCU"
   Button "HmiScreenItemData_2" at 1129,1 size 150x40; TextOn 'Back'; TextOff 'BWTS Setup'
      on Release: ActivateScreen("Balast Water Treatment Setup", 0)
   TextField "Text field_1" at 290,107 size 68x30; Text 'Tank Selected'
   TextField "Text field_2" at 841,107 size 61x30; Text 'BWTS Started'
   TextField "Text field_3" at 568,107 size 62x30; Text 'IGGS Started'
   TextField "Text field_4" at 659,107 size 60x30; Text 'GCU Started'
   TextField "Text field_5" at 748,107 size 61x30; Text 'PGC Started'
   TextField "Text field_6" at 908,107 size 102x30; Text 'Gas Transfer Started'
   Circle "Circle_10" at 956,89 size 14x14
      Appearance <- "2110_BTCS_CNTRL_DB_BTCS_STEP"
   TextField "Text field_7" at 995,107 size 125x30; Text 'Treatment Cycle Completed'
   TextField "Text field_23" at 261,291 size 34x14; Text 'MBG'
   GraphicView "Graphic view_17" at 575,446 size 532x12; Picture "Graphic_151"
   Button "Button_13" at 252,437 size 37x30; TextOff 'DB&B'
   TextField "Text field_58" at 188,226 size 50x40; Text 'Safe Area'
   Button "Button_20" at 724,152 size 115x34; TextOff 'Re-Oxygenation'
      Appearance <- "2110_BTCS_CNTRL_DB_BTCS_STEP"
   Button "Button_21" at 845,152 size 93x34; TextOff 'Post Dwell'
      Appearance <- "2110_BTCS_CNTRL_DB_BTCS_STATE"
   Circle "Circle_1" at 137,105 size 29x29
      Appearance <- "2110_BTCS_CNTRL_DB_BTCS_STATE"
   Circle "Circle_8" at 775,89 size 14x14
      Appearance <- "2110_BTCS_CNTRL_DB_BTCS_STEP"
   Circle "Circle_9" at 685,89 size 14x14
      Appearance <- "100_GCU_AUTO_SEQ_DB_CRNT_STEP"
   Circle "Circle_11" at 595,89 size 14x14
      Appearance <- "51_SLAVE_STATUS_RUNNING"
   Circle "Circle_12" at 866,89 size 14x14
      Appearance <- "2110_BTCS_CNTRL_DB_BTCS_STEP"
   Circle "Circle_13" at 324,89 size 14x14
      Appearance <- "HMI Indication Logic_DB_Tank Selected"
   Circle "Circle_14" at 414,89 size 14x14
      Appearance <- "2102_TIME_CALCS_DB_PRE_DWELL_TMR_DN"
   Button "Button_3" at 626,152 size 93x34; TextOff 'Dwell'
      Appearance <- "2110_BTCS_CNTRL_DB_BTCS_STATE"
   Button "Button_5" at 944,152 size 93x34; TextOff 'Complete'
      Appearance <- "HMI Indication Logic_DB_Sequence Finished"
   TextField "Text field_61" at 202,107 size 71x30; Text 'FA Mode Selected'
   Circle "Circle_2" at 230,89 size 14x14
      Appearance <- "HMI Indication Logic_DB_FA Mode Selected"
   TextField "Text field_60" at 190,519 size 46x25; Text 'GCU'
   GraphicIOField "Graphic I/O field_4" at 187,543 size 53x55; PictureList "GCU"
      ProcessValue <- "100_GCU_AUTO_SEQ_DB_RNG"
   TextField "Text field_74" at 186,279 size 54x25; Text 'IGGS'
   GraphicIOField "Graphic I/O field_1" at 185,303 size 57x53; PictureList "IGGS"
      ProcessValue <- "14_DQ_Data_24PF1"
   TextField "Text field_62" at 183,359 size 60x20; Text 'Disabled'
   TextField "Text field_77" at 183,359 size 60x20; Text 'Enabled'
      Visibility <- "51_SLAVE_STATUS_RUNNING"
   Button "Button_8" at 178,280 size 70x105; TextOff 'Text'
      on Release: ActivateScreen("Inert Gas Generator Plant", 0)
   TextField "Text field_70" at 183,599 size 60x20; Text 'Disabled'
   TextField "Text field_71" at 183,599 size 60x20; Text 'Enabled'
      Visibility <- "100_GCU_AUTO_SEQ_DB_RNG"
   Button "Button_4" at 178,521 size 70x105; TextOff 'Text'
      on Release: ActivateScreen("Inert Gas Conditioning Plant", 0)
   GraphicIOField "Graphic I/O field_2" at 770,45 size 250x30; PictureList "Process time Banner"
      Visibility <- "2110_BTCS_CNTRL_DB_BTCS_STATE"
      ProcessValue <- "2110_BTCS_CNTRL_DB_BTCS_STATE"
   Button "Button_14" at 303,152 size 93x34; TextOff 'Unselected'
      Visibility <- "HMI Indication Logic_DB_Tank Selected"
      Appearance <- "HMI Indication Logic_DB_Tank Selected"
   Button "Button_15" at 404,152 size 93x34; TextOff 'Selected'
      Appearance <- "HMI Indication Logic_DB_Tank Selected"
   Button "Button_16" at 506,152 size 115x34; TextOff 'De-Oxygenation'
      Appearance <- "2110_BTCS_CNTRL_DB_BTCS_STEP"
   TextField "Text field_92" at 304,351 size 76x15; Text 'FIT-418-6P'
   TextField "Text field_98" at 304,308 size 76x15; Text 'FIT-420-6P'
   Button "HmiScreenItemData_19" at 1185,676 size 72x27; TextOn 'Back'; TextOff 'Status'
      on Press: function_efd93a16("Treatment Status", 100, 471, -1, 3, 1)
   Group "Group_6" at 298,44 size 241x30
   Circle "Circle_26" at 504,89 size 14x14
      Appearance <- "2102_TIME_CALCS_DB_Time_To_Treatment"
   TextField "Text field_134" at 470,107 size 75x30; Text 'Wait for IGGS Start'
   GraphicView "Graphic view_4" at 357,210 size 25x62; Picture "Graphic_183"
   GraphicView "Graphic view_5" at 265,210 size 25x62; Picture "Graphic_183"
   IOField "I/O field_31" at 1053,45 size 225x30; FormatPattern ???????????????
      ProcessValue <- "Current User"
   Button "HmiScreenItemData_8" at 772,732 size 503x40; TextOn 'Back'; TextOff 'Text'